(* Logix 5000 project; controller PLC_MCC1300_75F1 vendor 1 type 14 code 166 rev 32.11; software revision 32.04; part 6 of 83 *)
(* tags used below, declared in another part *)
   M352 : MAC_Conveyor;
   M353 : MAC_Conveyor;
   N14 : DINT[500];
   N30 : DINT[32];
   N31 : DINT[33];   // M2 to M4
   N32 : DINT[33];
   N40 : DINT[32];
   N7 : DINT[101];
   N802 : INT[420];
   N803 : INT[420];
   O : INT[128];
   T4 : TIMER[51];
   T47 : TIMER[32];

ADD_ON_INSTRUCTION GP_TrackingGetLength   (* revision 1.0 *)
VAR_IN_OUT
   INO_tLine : UDT_LINE_TRACKING; {required}
END_VAR
VAR_INPUT
   IN_StartConveyorIndex : DINT; {access None, required}
   IN_StopConveyorIndex : DINT; {access None, required}
END_VAR
VAR_OUTPUT
   OUT_dLength_cmm : DINT; {access None}
END_VAR
VAR
   TMP_dLineSize : DINT; {access None}
   TMP_dIndex : DINT; {access None}
END_VAR

ROUTINE Logic   (* structured text *)
   
   OUT_dLength_cmm := 0;
   size(INO_tLine.rgtTrkConv[0],0,TMP_dLineSize);
   IF IN_StartConveyorIndex >= 0 AND IN_StartConveyorIndex < TMP_dLineSize AND IN_StopConveyorIndex >= IN_StartConveyorIndex AND IN_StopConveyorIndex < TMP_dLineSize THEN
   	FOR TMP_dIndex := IN_StartConveyorIndex TO IN_StopConveyorIndex DO
   		OUT_dLength_cmm := OUT_dLength_cmm + INO_tLine.rgtTrkConv[TMP_dIndex].dLengthConveyor;
   	END_FOR;
   END_IF;
   
END_ROUTINE
END_ADD_ON_INSTRUCTION

ADD_ON_INSTRUCTION GP_TrackingPresencePlate   (* revision 1.0 *)
VAR_INPUT
   IN_dPositionStartSearch_cmm : DINT; {access None, required}   // Position of start searching plate
   IN_dPositionStopSearch_cmm : DINT; {access None, required}   // Position of stop searching plate
   IN_xConvoySearchSingle : BOOL; {access None, required}   // Search single cap in a convoy
END_VAR
VAR_IN_OUT
   INO_tLine : UDT_LINE_TRACKING; {required}   // Tracking area
END_VAR
VAR_OUTPUT
   OUT_xPlatePresence : BOOL; {access Read Only, required}
END_VAR
VAR
   TMP_dIndConv : DINT; {access None}
   TMP_dPositionMax_cmm : DINT; {access None}
   TMP_dPositionMin_cmm : DINT; {access None}
   TMP_dIndConvMax : DINT; {access None}
   TMP_dIndConvMin : DINT; {access None}
   TMP_dIndCap : DINT; {access None}
   TMP_dLineSize : DINT; {access None}
END_VAR

ROUTINE Logic   (* structured text *)
   
   OUT_xPlatePresence := 0;
   TMP_dPositionMax_cmm := IN_dPositionStopSearch_cmm;
   TMP_dPositionMin_cmm := IN_dPositionStartSearch_cmm;
   size(INO_tLine.rgtTrkConv[0],0,TMP_dLineSize);
   
   //Search The index of Conveyor
   FOR TMP_dIndConv := 0 TO TMP_dLineSize - 1 DO
       //Search Conveyor Index Min
       IF TMP_dPositionMin_cmm <= INO_tLine.rgtTrkConv[TMP_dIndConv].dEndPosition_cmm AND TMP_dPositionMin_cmm >= INO_tLine.rgtTrkConv[TMP_dIndConv].dStartPosition_cmm THEN
           TMP_dIndConvMin := TMP_dIndConv;
       END_IF;
       //Search Conveyor Index Max
       IF TMP_dPositionMax_cmm <= INO_tLine.rgtTrkConv[TMP_dIndConv].dEndPosition_cmm AND TMP_dPositionMax_cmm >= INO_tLine.rgtTrkConv[TMP_dIndConv].dStartPosition_cmm THEN
           TMP_dIndConvMax := TMP_dIndConv;
           EXIT;
       END_IF;
   END_FOR;
   
   FOR TMP_dIndConv := TMP_dIndConvMin TO TMP_dIndConvMax DO
       IF INO_tLine.rgtTrkConv[TMP_dIndConv].xGlassPresence THEN
           FOR TMP_dIndCap := 0 TO INO_tLine.rgtTrkConv[TMP_dIndConv].dIndexCaps DO
               OUT_xPlatePresence := (INO_tLine.rgtTrkConv[TMP_dIndConv].Cap[TMP_dIndCap].dPresenceHead_cmm >= TMP_dPositionMin_cmm
   			AND INO_tLine.rgtTrkConv[TMP_dIndConv].Cap[TMP_dIndCap].dPresenceHead_cmm <= TMP_dPositionMax_cmm)
               OR (INO_tLine.rgtTrkConv[TMP_dIndConv].Cap[TMP_dIndCap].dPresenceTail_cmm >= TMP_dPositionMin_cmm
   			AND INO_tLine.rgtTrkConv[TMP_dIndConv].Cap[TMP_dIndCap].dPresenceTail_cmm <= TMP_dPositionMax_cmm)
   			OR (INO_tLine.rgtTrkConv[TMP_dIndConv].Cap[TMP_dIndCap].dPresenceHead_cmm >= TMP_dPositionMax_cmm
   			AND INO_tLine.rgtTrkConv[TMP_dIndConv].Cap[TMP_dIndCap].dPresenceTail_cmm <= TMP_dPositionMin_cmm);
               IF OUT_xPlatePresence THEN
                   EXIT;
               END_IF;
           END_FOR;
       END_IF;
       IF OUT_xPlatePresence THEN
           EXIT;
       END_IF;
   END_FOR;
   
END_ROUTINE
END_ADD_ON_INSTRUCTION

ADD_ON_INSTRUCTION GP_TrackingSearchIDPlate   (* revision 1.0 *)
VAR_IN_OUT
   INO_tBufferPlate : UDT_LINE_BUFFER_PLATE; {required}
END_VAR
VAR_INPUT
   IN_dIDPlate : DINT; {access None, required}
END_VAR
VAR_OUTPUT
   OUT_dIndexPlate : DINT; {access None, required}
   OUT_xPlateIDFound : BOOL; {access Read Only, required}
END_VAR
VAR_IN_OUT
   INO_CONST_dMaxLites : DINT; {constant, required}
   INO_CONST_dMaxCaps : DINT; {constant, required}
END_VAR
VAR
   TMP_dInd : DINT; {access None}
   TMP_dLite : DINT; {access None}
   TMP_dCap : DINT; {access None}
   TMP_dBufferSize : DINT; {access None}
END_VAR

ROUTINE Logic   (* structured text *)
   
   size(INO_tBufferPlate.rgtPlate[0],0,TMP_dBufferSize);
   OUT_dIndexPlate := 0;//reset Output
   //Search Plate Index
   IF IN_dIDPlate <> 0 THEN
       FOR TMP_dInd := 0 TO TMP_dBufferSize - 1 DO
           FOR TMP_dCap := 0 TO INO_CONST_dMaxCaps - 1 DO
               FOR TMP_dLite := 0 TO INO_CONST_dMaxLites - 1 DO
   				IF INO_tBufferPlate.rgtPlate[TMP_dInd].tData.rgtCap[TMP_dCap].rgtLite[TMP_dLite].dID = IN_dIDPlate THEN
   					OUT_xPlateIDFound := 1;
   				END_IF;
                   IF OUT_xPlateIDFound THEN
                       OUT_dIndexPlate := TMP_dInd;//When found plate Exit from function
                       TND( );
                   END_IF;
               END_FOR;
           END_FOR;
       END_FOR;
   END_IF;
   
END_ROUTINE
END_ADD_ON_INSTRUCTION

ADD_ON_INSTRUCTION GP_TrackingSearchPlate   (* revision 1.0 *)
VAR_INPUT
   IN_dPositionStartSearch_cmm : DINT; {access None, required}   // Position of start searching plate
   IN_dPositionStopSearch_cmm : DINT; {access None, required}   // Position of stop searching plate
   IN_xConvoySearchSingle : BOOL; {access None, required}   // Search single cap in a convoy
END_VAR
VAR_IN_OUT
   INO_tLineTracking : UDT_LINE_TRACKING; {required}   // Tracking area
   INO_GP_SearchPlate : GP_TrackingSearchPlate_STC; {required}   // Search results
   INO_dNumOfConveyors : DINT; {constant, required}   // Number of conveyors in tracking area
   INO_dNumCapsConveyor : DINT; {constant, required}   // Max number of caps per conveyor
   INO_tLineBufferPlate : UDT_LINE_BUFFER_PLATE; {required}   // Buffer plate
END_VAR
VAR
   TMP_dIndConv : DINT; {access None}
   TMP_dPositionMax_cmm : DINT; {access None}
   TMP_dPositionMin_cmm : DINT; {access None}
   TMP_xStartGreater : BOOL; {access None}
   TMP_dIndConvMax : DINT; {access None}
   TMP_dIndConvMin : DINT; {access None}
   TMP_dIndCap : DINT; {access None}
   TMP_dHeadPos : DINT; {access None}
   TMP_DIndexOut : DINT; {access None}
   TMP_dLastPosHead_cmm : DINT; {access None}
   TMP_dLastPosTail_cmm : DINT; {access None}
   TMP_dTailPos : DINT; {access None}
   TMP_dPointerCap : DINT; {access None}
   TMP_dTailPointer : DINT; {access None}
   TMP_dHeadPointer : DINT; {access None}   // Head pointer
END_VAR

ROUTINE Logic   (* structured text *)
   
   //Start Greater of the END
   TMP_xStartGreater := IN_dPositionStartSearch_cmm >= IN_dPositionStopSearch_cmm;
   INO_GP_SearchPlate.xTailPresence := 0;
   INO_GP_SearchPlate.xHeadPresence := 0;
   
   FOR TMP_DIndexOut := 0 TO 4 DO
       INO_GP_SearchPlate.rgdHead_cmm[TMP_DIndexOut] := 0;
       INO_GP_SearchPlate.rgdTail_cmm[TMP_DIndexOut] := 0;
       INO_GP_SearchPlate.rgdHeadPointer[TMP_DIndexOut] := 0;
       INO_GP_SearchPlate.rgdTailPointer[TMP_DIndexOut] := 0;
       INO_GP_SearchPlate.rgxHead.[TMP_DIndexOut] := 0;
       INO_GP_SearchPlate.rgxTail.[TMP_DIndexOut] := 0;
   END_FOR;
   TMP_DIndexOut := 0;
   
   IF TMP_xStartGreater THEN
       TMP_dPositionMax_cmm := IN_dPositionStartSearch_cmm;
       TMP_dPositionMin_cmm := IN_dPositionStopSearch_cmm;
   ELSE
       TMP_dPositionMax_cmm := IN_dPositionStopSearch_cmm;
       TMP_dPositionMin_cmm := IN_dPositionStartSearch_cmm;
   END_IF;
   
   //Search The index of Conveyor
   FOR TMP_dIndConv := 0 TO INO_dNumOfConveyors - 1 DO
       //Search Conveyor Index Min
       IF  TMP_dPositionMin_cmm <= INO_tLineTracking.rgtTrkConv[TMP_dIndConv].dEndPosition_cmm
   		AND TMP_dPositionMin_cmm >= INO_tLineTracking.rgtTrkConv[TMP_dIndConv].dStartPosition_cmm THEN
           TMP_dIndConvMin := TMP_dIndConv;
       END_IF;
       //Search Conveyor Index Max
       IF TMP_dPositionMax_cmm <= INO_tLineTracking.rgtTrkConv[TMP_dIndConv].dEndPosition_cmm
   		AND TMP_dPositionMax_cmm >= INO_tLineTracking.rgtTrkConv[TMP_dIndConv].dStartPosition_cmm THEN
           TMP_dIndConvMax := TMP_dIndConv;
           EXIT;
       END_IF;
   END_FOR;
   
   IF TMP_xStartGreater THEN
       //Start To the Max
   
       TMP_dLastPosHead_cmm := TMP_dPositionMax_cmm+1;
       TMP_dLastPosTail_cmm := TMP_dPositionMax_cmm+1;
       FOR TMP_DIndexOut := 0 TO 4 DO
           TMP_dHeadPos := 0;
           TMP_dTailPos := 0;
           FOR TMP_dIndConv := TMP_dIndConvMax TO TMP_dIndConvMin BY -1 DO
               IF INO_tLineTracking.rgtTrkConv[TMP_dIndConv].xGlassPresence THEN
                   FOR TMP_dIndCap := 0 TO INO_tLineTracking.rgtTrkConv[TMP_dIndConv].dIndexCaps DO
   					IF TMP_dIndCap < INO_dNumCapsConveyor THEN //Check to avoid CPU fault in case of tracking errors
   	                    TMP_dPointerCap := INO_tLineTracking.rgtTrkConv[TMP_dIndConv].Cap[TMP_dIndCap].dPointer;
   	                    IF INO_tLineTracking.rgtTrkConv[TMP_dIndConv].Cap[TMP_dIndCap].dHeadPos_cmm >= TMP_dPositionMin_cmm
   	                        AND INO_tLineTracking.rgtTrkConv[TMP_dIndConv].Cap[TMP_dIndCap].dHeadPos_cmm <= TMP_dPositionMax_cmm
   							AND INO_tLineTracking.rgtTrkConv[TMP_dIndConv].Cap[TMP_dIndCap].dHeadPos_cmm >= TMP_dHeadPos
   	                        AND (INO_tLineBufferPlate.rgtPlate[TMP_dPointerCap].tTracking.dPreviousCapIndex <= 0 OR IN_xConvoySearchSingle)
   							AND INO_tLineTracking.rgtTrkConv[TMP_dIndConv].Cap[TMP_dIndCap].xHead
   	                        AND INO_tLineTracking.rgtTrkConv[TMP_dIndConv].Cap[TMP_dIndCap].dHeadPos_cmm < TMP_dLastPosHead_cmm
   	                        AND ((NOT INO_tLineBufferPlate.rgtPlate[TMP_dPointerCap].tTracking.xNotConsConvTrk)
   							OR TMP_dIndConv < INO_tLineBufferPlate.rgtPlate[TMP_dPointerCap].tTracking.dIndexConvNotCons) THEN
   	                        TMP_dHeadPos := INO_tLineTracking.rgtTrkConv[TMP_dIndConv].Cap[TMP_dIndCap].dHeadPos_cmm;
   	                        TMP_dHeadPointer := TMP_dPointerCap;
   	                    END_IF;
   
   	                    IF INO_tLineTracking.rgtTrkConv[TMP_dIndConv].Cap[TMP_dIndCap].dTailPos_cmm >= TMP_dPositionMin_cmm
   	                        AND INO_tLineTracking.rgtTrkConv[TMP_dIndConv].Cap[TMP_dIndCap].dTailPos_cmm <= TMP_dPositionMax_cmm
   							AND INO_tLineTracking.rgtTrkConv[TMP_dIndConv].Cap[TMP_dIndCap].dTailPos_cmm >= TMP_dTailPos
   	                        AND (INO_tLineBufferPlate.rgtPlate[TMP_dPointerCap].tTracking.dNextCapIndex <= 0
   							OR IN_xConvoySearchSingle) AND INO_tLineTracking.rgtTrkConv[TMP_dIndConv].Cap[TMP_dIndCap].xTail
   	                        AND INO_tLineTracking.rgtTrkConv[TMP_dIndConv].Cap[TMP_dIndCap].dTailPos_cmm < TMP_dLastPosTail_cmm
   	                        AND ((NOT INO_tLineBufferPlate.rgtPlate[TMP_dPointerCap].tTracking.xNotConsConvTrk)
   							OR TMP_dIndConv < INO_tLineBufferPlate.rgtPlate[TMP_dPointerCap].tTracking.dIndexConvNotCons) THEN
   	                        TMP_dTailPos := INO_tLineTracking.rgtTrkConv[TMP_dIndConv].Cap[TMP_dIndCap].dTailPos_cmm;
   	                        TMP_dTailPointer := TMP_dPointerCap;
   	                    END_IF;
   					END_IF;
                   END_FOR;
               END_IF;
           END_FOR;
           //Write Output
           IF TMP_dHeadPointer <> 0 THEN
               INO_GP_SearchPlate.rgdHead_cmm[TMP_DIndexOut] := TMP_dHeadPos;
               INO_GP_SearchPlate.rgdHeadPointer[TMP_DIndexOut] := TMP_dHeadPointer;
               INO_GP_SearchPlate.rgxHead.[TMP_DIndexOut] := 1;
               INO_GP_SearchPlate.xHeadPresence := 1;
               TMP_dLastPosHead_cmm := TMP_dHeadPos;
               TMP_dHeadPointer := 0;
           END_IF;
   
           IF TMP_dTailPointer <> 0 THEN
               INO_GP_SearchPlate.rgdTail_cmm[TMP_DIndexOut] := TMP_dTailPos;
               INO_GP_SearchPlate.rgdTailPointer[TMP_DIndexOut] := TMP_dTailPointer;
               INO_GP_SearchPlate.rgxTail.[TMP_DIndexOut] := 1;
               INO_GP_SearchPlate.xTailPresence := 1;
               TMP_dLastPosTail_cmm := TMP_dTailPos;
           END_IF;
   
           IF TMP_dTailPointer = 0 AND TMP_dHeadPointer = 0 THEN
               EXIT;
           END_IF;
           TMP_dTailPointer := 0;
           TMP_dHeadPointer := 0;
       END_FOR;
   
   ELSE
       TMP_dLastPosHead_cmm := TMP_dPositionMin_cmm - 1;
       TMP_dLastPosTail_cmm := TMP_dPositionMin_cmm - 1;
       //Start To the Min
       FOR TMP_DIndexOut := 0 TO 4 DO
           TMP_dHeadPos := TMP_dPositionMax_cmm;
           TMP_dTailPos := TMP_dPositionMax_cmm;
           FOR TMP_dIndConv := TMP_dIndConvMin TO TMP_dIndConvMax DO
   
               IF INO_tLineTracking.rgtTrkConv[TMP_dIndConv].xGlassPresence THEN
                   FOR TMP_dIndCap := 0 TO INO_tLineTracking.rgtTrkConv[TMP_dIndConv].dIndexCaps DO
   					IF TMP_dIndCap < INO_dNumCapsConveyor THEN // To avoid CPU fault in case of tracking error (too much caps in one conveyor)
   	                    TMP_dPointerCap := INO_tLineTracking.rgtTrkConv[TMP_dIndConv].Cap[TMP_dIndCap].dPointer;
   	                    IF INO_tLineTracking.rgtTrkConv[TMP_dIndConv].Cap[TMP_dIndCap].dHeadPos_cmm >= TMP_dPositionMin_cmm
   	                        AND INO_tLineTracking.rgtTrkConv[TMP_dIndConv].Cap[TMP_dIndCap].dHeadPos_cmm <= TMP_dPositionMax_cmm
   							AND INO_tLineTracking.rgtTrkConv[TMP_dIndConv].Cap[TMP_dIndCap].dHeadPos_cmm <= TMP_dHeadPos
   	                        AND (INO_tLineBufferPlate.rgtPlate[TMP_dPointerCap].tTracking.dPreviousCapIndex <= 0 OR IN_xConvoySearchSingle)
   							AND INO_tLineTracking.rgtTrkConv[TMP_dIndConv].Cap[TMP_dIndCap].xHead
   	                        AND INO_tLineTracking.rgtTrkConv[TMP_dIndConv].Cap[TMP_dIndCap].dHeadPos_cmm > TMP_dLastPosHead_cmm THEN
   	                        TMP_dHeadPos := INO_tLineTracking.rgtTrkConv[TMP_dIndConv].Cap[TMP_dIndCap].dHeadPos_cmm;
   	                        TMP_dHeadPointer := TMP_dPointerCap;
   	                    END_IF;
   
   	                    IF INO_tLineTracking.rgtTrkConv[TMP_dIndConv].Cap[TMP_dIndCap].dTailPos_cmm >= TMP_dPositionMin_cmm
   	                        AND INO_tLineTracking.rgtTrkConv[TMP_dIndConv].Cap[TMP_dIndCap].dTailPos_cmm <= TMP_dPositionMax_cmm
   							AND INO_tLineTracking.rgtTrkConv[TMP_dIndConv].Cap[TMP_dIndCap].dTailPos_cmm <= TMP_dTailPos
   	                        AND (INO_tLineBufferPlate.rgtPlate[TMP_dPointerCap].tTracking.dNextCapIndex <= 0 OR IN_xConvoySearchSingle)
   							AND INO_tLineTracking.rgtTrkConv[TMP_dIndConv].Cap[TMP_dIndCap].xTail
   	                        AND INO_tLineTracking.rgtTrkConv[TMP_dIndConv].Cap[TMP_dIndCap].dTailPos_cmm > TMP_dLastPosTail_cmm THEN
   	                        TMP_dTailPos := INO_tLineTracking.rgtTrkConv[TMP_dIndConv].Cap[TMP_dIndCap].dTailPos_cmm;
   	                        TMP_dTailPointer := TMP_dPointerCap;
   	                    END_IF;
   					END_IF;
   	            END_FOR;
               END_IF;
           END_FOR;
           //Write Output
           IF TMP_dHeadPointer <> 0 THEN
               INO_GP_SearchPlate.rgdHead_cmm[TMP_DIndexOut] := TMP_dHeadPos;
               INO_GP_SearchPlate.rgdHeadPointer[TMP_DIndexOut] := TMP_dHeadPointer;
               INO_GP_SearchPlate.rgxHead.[TMP_DIndexOut] := 1;
               INO_GP_SearchPlate.xHeadPresence := 1;
               TMP_dLastPosHead_cmm := TMP_dHeadPos;
               TMP_dHeadPointer := 0;
           END_IF;
   
           IF TMP_dTailPointer <> 0 THEN
               INO_GP_SearchPlate.rgdTail_cmm[TMP_DIndexOut] := TMP_dTailPos;
               INO_GP_SearchPlate.rgdTailPointer[TMP_DIndexOut] := TMP_dTailPointer;
               INO_GP_SearchPlate.rgxTail.[TMP_DIndexOut] := 1;
               INO_GP_SearchPlate.xTailPresence := 1;
               TMP_dLastPosTail_cmm := TMP_dTailPos;
           END_IF;
   
           IF TMP_dTailPointer = 0 AND TMP_dHeadPointer = 0 THEN
               EXIT;
           END_IF;
           TMP_dTailPointer := 0;
           TMP_dHeadPointer := 0;
       END_FOR;
   END_IF;
   
END_ROUTINE
END_ADD_ON_INSTRUCTION

ADD_ON_INSTRUCTION GP_TrackingValidateIndex   (* revision 1.0 *)
VAR_IN_OUT
   INO_tLineBufferPlate : UDT_LINE_BUFFER_PLATE; {required}   // Buffer Plate
   INO_dIDMemory : DINT; {required}   // Memory of ID
END_VAR
VAR_INPUT
   IN_dIndex : DINT; {access None, required}   // Index
END_VAR
VAR_OUTPUT
   OUT_xDataConsistance : BOOL; {access None, required}   // Data consistance
END_VAR

ROUTINE Logic   (* structured text *)
   
   IF IN_dIndex <> 0 THEN
   	IF INO_tLineBufferPlate.rgtPlate[IN_dIndex].tData.rgtCap[0].dID <> 0 AND (INO_tLineBufferPlate.rgtPlate[IN_dIndex].tData.rgtCap[0].dID = INO_dIDMemory OR INO_dIDMemory = 0) THEN
   		OUT_xDataConsistance := 1;
   	ELSE
   		OUT_xDataConsistance := 0;
   		INO_dIDMemory := 0;
   	END_IF;
   ELSE
   	INO_dIDMemory := 0;
   	OUT_xDataConsistance := 0;
   END_IF;
   
END_ROUTINE
END_ADD_ON_INSTRUCTION

VAR_GLOBAL   (* controller tags *)
   AUX_tBufferPlate_NULL : UDT_BufferPlate; {access Read Only}
   AUX_tCapsConveyor_NULL : UDT_CapsConveyor_ZC; {access Read Only}
   AUX_tConvoy_SL_NULL : UDT_Convoy_SL; {access Read Only}
   AUX_tConvoyCap_ZC_NULL : UDT_ConvoyCap_ZC; {access Read Only}
   AUX_tHMI_Lite_NULL : UDT_HMI_LITE; {access Read Only}
   AUX_xDebugNewPlate : BOOL; {access Read Only}
   AUX_xInitialize : BOOL; {access Read Only}
   Axies : MOTION_GROUP; {access Read Only}
   B102 : DINT[1];
   B107 : DINT[1];
   B112 : DINT[1];
   B117 : DINT[1];
   B122 : DINT[1];
   B127 : DINT[1];
   B132 : DINT[1];
   B151 : DINT[1];
   B152 : DINT[1];
   B153 : DINT[1];
   B154 : DINT[1];
   B155 : DINT[1];
   B156 : DINT[1];
   B157 : DINT[1];
   B158 : DINT[1];
   B159 : DINT[1];
   B160 : DINT[1];
   B161 : DINT[1];
   B162 : DINT[1];
   B163 : DINT[1];
   B164 : DINT[1];
   B165 : DINT[1];
   B166 : DINT[1];
   B167 : DINT[1];
   B168 : DINT[1];
   B169 : DINT[1];
   B170 : DINT[1];
   B171 : DINT[1];
   B172 : DINT[1];
   B175 : DINT[1];
   B176 : DINT[1] := ([0] := 2#0000_0000_0000_0000_0000_1100_0000_0000);
   B180 : DINT[10] := ([0] := 2#0000_0000_0000_0000_0001_1111_1001_0000, [1] := 2#0000_0000_0000_0000_0000_0000_0000_0001, [2] := 2#0000_0000_0000_0000_0001_0000_1011_0111, [4] := 2#0000_0000_0000_0000_0001_0000_0000_0000, [5] := 2#0000_0000_0000_0000_0000_0000_0011_0001, [6] := 2#0000_0000_0000_0000_1001_1110_0000_0000, [7] := 2#0000_0000_0000_0000_0001_0110_1101_1011, [9] := 2#0000_0000_0000_0000_0000_0000_1100_0000);
   B3 : DINT[51] := ([0] := 2#0000_0000_0000_0000_0010_0000_0000_0000, [1] := 2#0000_0000_0000_0000_0000_0000_1000_0000, [6] := 2#0000_0000_0000_0000_0000_0010_0000_0000, [7] := 2#0000_0000_0000_0000_1000_0000_0000_1000, [50] := 2#0000_0000_0000_0000_0000_0000_0001_0000);
        [0].0   // DUMMY for Red Stack lite
        [0].1   // VMCC M4 Mainline is Backed up Flush a CAP
        [10].14   // Always false Tony
        [10].15   // Tony test Bit
        [12].12   // M3CM04 Second. Trans. Conv 4 - Resync Photo-Eye North (Conveyor 4)
        [12].13   // M3CM05 Second. Trans. Conv 5 - Resync Photo-Eye North (Conveyor 5)
        [12].14   // M3CM06 Second. Trans. Conv 6 - Resync Photo-Eye North (Conveyor 6)
        [12].15   // M3CM07 Queue Conv 2 Resync Photo-Eye North (Conveyor 7)
        [13].0   // M3CM08 Queue Conv 3 Resync Photo-Eye North (Conveyor 8)
        [13].1   // M3CM08 Queue Conv 4 Resync Photo-Eye North (Conveyor 9)
        [13].2   // QUALITY SAMPLE XFER 201.010 Xfer Conv M3CM10 QC5 Resync PE North (Conveyor 10)
        [13].6   // TRANSFER 1A VHSC gating Photo-eye North
        [14].0   // Mainline is in Sleep Mode
        [14].1   // Mainline in Sleep Mode Stop Conveyors
        [14].2   // ink jet ons
        [14].3   // INK JET Cap needs Ink jet messg
        [14].4   // ink jet ons2
        [18].13   // TRANSFER 1 Oversize cap Photo-eye EAST
        [18].14   // TRANSFER 1 Oversize cap Photo-Eye WEST
        [18].15   // TRANSFER 1A Oversize cap Photo-eye EAST
        [19].0   // TRANSFER 1A Oversize cap Photo-Eye WEST
        [2].15   // M4 -->> M5 Cap information One shot
        [50].0   // Sample Shuttle Peg is Approaching
        [50].1   // Sample Shuttle Peg is Ready for Pick up
        [5].10   // VMCC 4 Drive Fault Has occurred
        [5].11   // VMCC 3 Drive fault Has occurred
        [6].10   // CONVEYOR 6 Resync Photo-Eye South M3CM06
        [6].11   // M3CM07 Queue Conv 2 Resync Photo-Eye South (Conveyor 7)
        [6].12   // M3CM08 Queue Conv 3 Resync Photo-Eye South (Conveyor 8)
        [6].13   // M3CM08 Queue Conv 4 Resync Photo-Eyes (Conveyor 9)
        [6].14   // QUALITY SAMPLE XFER 201.010 Xfer Conv M3CM10 QC 5 Resync PE South (Conveyor 10)
        [6].15   // M4CM04 Transfer 1 Resync Photo-Eye South (Conveyor 11)
        [6].8   // M3CM04 Second. Trans. Conv 4 - Resync Photo-Eye South (Conveyor 4)
        [6].9   // M3CM05 Second. Trans. Conv 5 - Resync Photo-Eye South (Conveyor 5)
        [7].0   // M4CM03 Transfer 1 Rolls B Resync Photo-Eye South (Conveyor 12)
        [7].1   // M4CM04 Transfer 1 Rolls C Resync Photo-Eye South (Conveyor 13)
        [7].2   // TRANSFER 1A VHSC gating Photo-eye South
        [7].3   // M4CM05 Transfer 1A Rolls A - Rsync Photo-Eye South (Conveyor 15)
        [7].4   // M4CM07 Transfer 1A Rolls B - Rsync Photo-Eye South (Conveyor 16)
        [7].5   // M4CM09 Transfer 1A Rolls C - Rsync Photo-Eye South (Conveyor 17)
   B41 : DINT[3] := ([2] := 2#0000_0000_0000_0000_1000_0000_0000_0000);
        [0].13   // Conveyor 13 Resync Window
        [0].14   // Conveyor 14 Resync Window
        [0].15   // Conveyor 15 Resync Window
        [0].2   // Conveyor 2 Resync Window
        [0].3   // Conveyor 3 Resync Window
        [0].4   // Conveyor 4 Resync Window
        [0].5   // Conveyor 5 Resync Window
        [0].6   // Conveyor 6 Resync Window
        [0].7   // Conveyor 7 Resync Window
        [0].8   // Conveyor 8 Resync Window
        [0].9   // Conveyor 9 Resync Window
        [1].0   // Conveyor 16 Resync Window
        [1].5   // Conveyor 21 Resync Window
        [1].6   // Conveyor 22 Resync Window
        [1].7   // Conveyor 23 Resync Window
        [1].8   // Conveyor 24 Resync Window
        [1].9   // Conveyor 25 Resync Window
        [2].0   // Conveyor 32 Resync Window
        [1].1   // Conveyor 17 Resync Window
        [1].10   // Conveyor 26 Resync Window
        [1].11   // Conveyor 27 Resync Window
        [1].12   // Conveyor 28 Resync Window
        [1].13   // Conveyor 29 Resync Window
        [1].14   // Conveyor 30 Resync Window
        [1].15   // Conveyor 31 Resync Window
        [1].2   // Conveyor 18 Resync Window
        [1].3   // Conveyor 19 Resync Window
        [1].4   // Conveyor 20 Resync Window
        [0].1   // Conveyor 1 Resync Window
        [0].10   // Conveyor 10 Resync Window
        [0].11   // Conveyor 11 Resync Window
        [0].12   // Conveyor 12 Resync Window
   B42 : DINT[3];
        [0].1   // Conveyor 1 Resync Input
        [0].10   // Conveyor 10 Resync Input
        [0].11   // Conveyor 11 Resync Input
        [0].12   // Conveyor 12 Resync Input
        [0].13   // Conveyor 13 Resync Input
        [0].14   // Conveyor 14 Resync Input
        [0].15   // Conveyor 15 Resync Input
        [0].2   // Conveyor 2 Resync Input
        [0].3   // Conveyor 3 Resync Input
        [0].4   // Conveyor 4 Resync Input
        [0].5   // Conveyor 5 Resync Input
        [0].6   // Conveyor 6 Resync Input
        [0].7   // Conveyor 7 Resync Input
        [0].8   // Conveyor 8 Resync Input
        [0].9   // Conveyor 9 Resync Input
        [1].0   // Conveyor 16 Resync Input
        [1].1   // Conveyor 17 Resync Input
        [1].10   // Conveyor 26 Resync Input
        [1].11   // Conveyor 27 Resync Input
        [1].12   // Conveyor 28 Resync Input
        [1].13   // Conveyor 29 Resync Input
        [1].14   // Conveyor 30 Resync Input
        [1].15   // Conveyor 31 Resync Input
        [1].2   // Conveyor 18 Resync Input
        [1].3   // Conveyor 19 Resync Input
        [1].4   // Conveyor 20 Resync Input
        [1].5   // Conveyor 21 Resync Input
        [1].6   // Conveyor 22 Resync Input
        [1].7   // Conveyor 23 Resync Input
        [1].8   // Conveyor 24 Resync Input
        [1].9   // Conveyor 25 Resync Input
        [2].0   // Conveyor 32 Resync Input
   B43 : DINT[3];
        [0].12   // Conveyor 12 Resync Output
        [0].13   // Conveyor 13 Resync Output
        [0].14   // Conveyor 14 Resync Output
        [0].15   // Conveyor 15 Resync Output
        [0].2   // Conveyor 2 Resync Output
        [0].3   // Conveyor 3 Resync Output
        [0].4   // Conveyor 4 Resync Output
        [0].5   // Conveyor 5 Resync Output
        [0].6   // Conveyor 6 Resync Output
        [0].7   // Conveyor 7 Resync Output
        [0].8   // Conveyor 8 Resync Output
        [0].9   // Conveyor 9 Resync Output
        [1].0   // Conveyor 16 Resync Output
        [1].1   // Conveyor 17 Resync Output
        [1].10   // Conveyor 26 Resync Output
        [1].11   // Conveyor 27 Resync Output
        [1].12   // Conveyor 28 Resync Output
        [1].13   // Conveyor 29 Resync Output
        [1].14   // Conveyor 30 Resync Output
        [1].15   // Conveyor 31 Resync Output
        [1].2   // Conveyor 18 Resync Output
        [1].3   // Conveyor 19 Resync Output
        [1].4   // Conveyor 20 Resync Output
        [1].5   // Conveyor 21 Resync Output
        [1].6   // Conveyor 22 Resync Output
        [1].7   // Conveyor 23 Resync Output
        [1].8   // Conveyor 24 Resync Output
        [1].9   // Conveyor 25 Resync Output
        [2].0   // Conveyor 32 Resync Output
        [0].1   // Conveyor 1 Resync Output
        [0].10   // Conveyor 10 Resync Output
        [0].11   // Conveyor 11 Resync Output
   B45 : DINT[3];
        [0].13   // Conveyor 13 Resync Input Leading Edge
        [0].14   // Conveyor 14 Resync Input Leading Edge
        [0].15   // Conveyor 15 Resync Input Leading Edge
        [0].2   // Conveyor 2 Resync Input Leading Edge
        [0].3   // Conveyor 3 Resync Input Leading Edge
        [0].4   // Conveyor 4 Resync Input Leading Edge
        [0].5   // Conveyor 5 Resync Input Leading Edge
        [0].6   // Conveyor 6 Resync Input Leading Edge
        [0].7   // Conveyor 7 Resync Input Leading Edge
        [0].8   // Conveyor 8 Resync Input Leading Edge
        [0].9   // Conveyor 9 Resync Input Leading Edge
        [1].0   // Conveyor 16 Resync Input Leading Edge
        [1].1   // Conveyor 17 Resync Input Leading Edge
        [1].10   // Conveyor 26 Resync Input Leading Edge
        [1].11   // Conveyor 27 Resync Input Leading Edge
        [1].12   // Conveyor 28 Resync Input Leading Edge
        [1].13   // Conveyor 29 Resync Input Leading Edge
        [1].14   // Conveyor 30 Resync Input Leading Edge
        [1].15   // Conveyor 31 Resync Input Leading Edge
        [1].2   // Conveyor 18 Resync Input Leading Edge
        [1].3   // Conveyor 19 Resync Input Leading Edge
        [1].4   // Conveyor 20 Resync Input Leading Edge
        [1].5   // Conveyor 21 Resync Input Leading Edge
        [1].6   // Conveyor 22 Resync Input Leading Edge
        [1].7   // Conveyor 23 Resync Input Leading Edge
        [1].8   // Conveyor 24 Resync Input Leading Edge
        [1].9   // Conveyor 25 Resync Input Leading Edge
        [2].0   // Conveyor 32 Resync Input Leading Edge
        [0].1   // Conveyor 1 Resync Input Leading Edge
        [0].10   // Conveyor 10 Resync Input Leading Edge
        [0].11   // Conveyor 11 Resync Input Leading Edge
        [0].12   // Conveyor 12 Resync Input Leading Edge
   B46 : DINT[3];
        [1].11   // Conveyor 27 Resync Input Trailing Edge
        [0].1   // Conveyor 1 Resync Input Trailing Edge
        [1].12   // Conveyor 28 Resync Input Trailing Edge
        [1].13   // Conveyor 29 Resync Input Trailing Edge
        [0].10   // Conveyor 10 Resync Input Trailing Edge
        [1].14   // Conveyor 30 Resync Input Trailing Edge
        [1].15   // Conveyor 31 Resync Input Trailing Edge
        [0].11   // Conveyor 11 Resync Input Trailing Edge
        [1].2   // Conveyor 18 Resync Input Trailing Edge
        [1].3   // Conveyor 19 Resync Input Trailing Edge
        [0].12   // Conveyor 12 Resync Input Trailing Edge
        [1].4   // Conveyor 20 Resync Input Trailing Edge
        [1].5   // Conveyor 21 Resync Input Trailing Edge
        [0].13   // Conveyor 13 Resync Input Trailing Edge
        [1].6   // Conveyor 22 Resync Input Trailing Edge
        [0].14   // Conveyor 14 Resync Input Trailing Edge
        [0].15   // Conveyor 15 Resync Input Trailing Edge
        [1].7   // Conveyor 23 Resync Input Trailing Edge
        [0].2   // Conveyor 2 Resync Input Trailing Edge
        [1].8   // Conveyor 24 Resync Input Trailing Edge
        [1].9   // Conveyor 25 Resync Input Trailing Edge
        [0].3   // Conveyor 3 Resync Input Trailing Edge
        [0].4   // Conveyor 4 Resync Input Trailing Edge
        [0].5   // Conveyor 5 Resync Input Trailing Edge
        [0].6   // Conveyor 6 Resync Input Trailing Edge
        [0].7   // Conveyor 7 Resync Input Trailing Edge
        [0].8   // Conveyor 8 Resync Input Trailing Edge
        [0].9   // Conveyor 9 Resync Input Trailing Edge
        [2].0   // Conveyor 32 Resync Input Trailing Edge
        [1].0   // Conveyor 16 Resync Input Trailing Edge
        [1].1   // Conveyor 17 Resync Input Trailing Edge
        [1].10   // Conveyor 26 Resync Input Trailing Edge
   B60 : DINT[4];
        [0].12   // Conveyor 12 Glass in Transit Bits
        [0].13   // Conveyor 13 Glass in Transit Bits
        [0].14   // Conveyor 14 Glass in Transit Bits
        [0].15   // Conveyor 15 Glass in Transit Bits
        [0].2   // Conveyor 2 Glass in Transit Bits
        [0].3   // Conveyor 3 Glass in Transit Bits
        [0].4   // Conveyor 4 Glass in Transit Bits
        [0].5   // Conveyor 5 Glass in Transit Bits
        [0].6   // Conveyor 6 Glass in Transit Bits
        [0].7   // Conveyor 7 Glass in Transit Bits
        [0].8   // Conveyor 8 Glass in Transit Bits
        [0].9   // Conveyor 9 Glass in Transit Bits
        [1].0   // Conveyor 16 Glass in Transit Bits
        [1].1   // Conveyor 17 Glass in Transit Bits
        [1].10   // Conveyor 26 Glass in Transit Bits
        [1].11   // Conveyor 27 Glass in Transit Bits
        [1].12   // Conveyor 28 Glass in Transit Bits
        [1].13   // Conveyor 29 Glass in Transit Bits
        [1].14   // Conveyor 30 Glass in Transit Bits
        [1].15   // Conveyor 31 Glass in Transit Bits
        [1].2   // Conveyor 18 Glass in Transit Bits
        [1].3   // Conveyor 19 Glass in Transit Bits
        [1].4   // Conveyor 20 Glass in Transit Bits
        [1].5   // Conveyor 21 Glass in Transit Bits
        [1].6   // Conveyor 22 Glass in Transit Bits
        [1].7   // Conveyor 23 Glass in Transit Bits
        [1].8   // Conveyor 24 Glass in Transit Bits
        [0].1   // Conveyor 1 Glass in Transit Bits
        [1].9   // Conveyor 25 Glass in Transit Bits
        [0].10   // Conveyor 10 Glass in Transit Bits
        [0].11   // Conveyor 11 Glass in Transit Bits
        [2].0   // Conveyor 32 Glass in Transit Bits
   B70 : DINT[13] := ([4] := 2#0000_0000_0000_0000_0000_0000_0000_0010, [6] := 2#0000_0000_0000_0000_0100_0000_0000_0000, [8] := 2#0000_0000_0000_0000_1101_0000_0000_1100);
        [0]   // TRANSFER 1 Status Bits
        [0].0   // TRANSFER 1 One conveyor transfer
        [0].1   // TRANSFER 1 Downstream half of transfer occuppied
        [0].2   // TRANSFER 1 Two conveyor Transfer
        [0].3   // TRANSFER 1 Downstream Total transfer Occupied
        [0].4   // TRANSFER 1 Three conveyor Transfer
        [0].5   // TRANSFER 1 Sample plate for Transfer 1
        [1].12   // TRANSFER 1 Upstream Cap is stopped at transfer
        [1].13   // TRANSFER 1 Downstream Cap is stopped at transfer
        [1].2   // TRANSFER 1 Lash Rolls A to Rolls B (i.e. force them to follow)
        [1].4   // TRANSFER 1 Upstream half of transfer Wait to see Gate input
        [1].5   // TRANSFER 1 Downstream half of transfer Wait to see Gate Input
        [1].8   // TRANSFER 1 Upstream half of Transfer VHSC Control Enabled
        [1].9   // TRANSFER 1 Downstream Half of Transfer VHSC Control Enabled
        [3].11   // TRANSFER 1 Leading cap Has exited xfer On upstream half only xfer
        [3].12   // TRANSFER 1 Trail edge Lock input
        [3].13   // TRANSFER 1 Conveyor is Seized for Transfer
        [4].0   // TRANSFER 1 Flush Signal
        [4].1   // TRANSFER 1 Setup Subroutine Glass Must Be Rotated before Packing
        [4].10   // TRANSFER 1 Rolls B Resync window Is a Two-Conv Transfer Cap
        [4].14   // TRANSFER 1 Glass was Aborted O/S
        [4].15   // TRANSFER 1 Occupied or Positioning a Cap
        [4].6   // TRANSFER 1 Transfer ABORTED!
        [4].7   // TRANSFER 1 Transfer is Complete
        [4].9   // TRANSFER 1 Stream 1 Size Matches the Jumbo Setup Size
        [5].1   // TRANSFER 1 Oversize cap Stopped at Transfer
        [5].15   // TRANSFER 1 Deck has been Raised manually
        [5].2   // TRANSFER 1 Glass is Ready for Transfer & No Vision Results Received when needed
        [5].3   // TRANSFER 1 Glass is Ready for Transfer & Vision Results were Received
        [6]   // TRANSFER 1 Transfer abort Reason History Bits
        [6].0   // Transfer abort Reason History Bit MANUAL ABORT
        [6].1   // REASON 1 Transfer Abort - Rack fault
        [6].10   // REASON 10 Transfer Abort - Deck raise Failure
        [6].11   // REASON 11 Transfer Abort - Duration Watchdog
        [6].12   // REASON 12 Transfer Abort - Size Mismatch
        [6].13   // REASON 13 Transfer Abort - Mainline Flush
        [6].14   // REASON 14 Transfer Abort - Transfer Disable Switch
        [6].15   // REASON 15 Transfer Abort - Mainline Vision Reject
        [6].2   // REASON 2 Transfer Abort - Leg equip. Failure
        [6].3   // REASON 3 Transfer Abort - Bad cap data To leg PLC
        [6].4   // REASON 4 Transfer Abort - Belt drive Fault
        [6].5   // REASON 5 Transfer Abort - LCR watchdog
        [6].6   // REASON 6 Transfer Abort - Rolls A Stop Watchdog
        [6].7   // REASON 7 Transfer Abort - Rolls B Stop Watchdog
        [6].8   // REASON 8 Transfer Abort - Rolls A Oversize cap
        [6].9   // REASON 9 Transfer Abort - Rolls B Oversize cap
        [7].0   // TRANSFER 1 One conveyor LCR
        [7].1   // TRANSFER 1 Downstream half Transfer LCR
        [7].2   // TRANSFER 1 Two conveyor LCR
        [7].3   // TRANSFER 1 Downstream Full Size Transfer LCR
        [7].4   // TRANSFER 1 Three conveyor LCR
        [8].0   // TRANSFER 1 Leading Cap Runout In Progress
        [8].1   // TRANSFER 1 Gap too small For one Conveyor Transfer
        [8].12   // TRANSFER 1 Conveyor 6 run permissives
        [8].13   // TRANSFER 1 Cap at Photo-Eye will Resync
        [8].15   // Valid data
        [8].2   // TRANSFER 1 Gap too small For two Conveyor Transfer
        [8].3   // TRANSFER 1 Gap too small For three Conveyor Transfer
        [8].4   // TRANSFER 1 Minimum gap For DECEL Is not Present!
        [9].0   // TRANSFER 1 Runout Sensors Checked OK Reset Warning Seal Circuit
        [9].1   // TRANSFER 1 Glass is Long enough to Reach the Center Runout Sensor
        [9].2   // TRANSFER 1 Glass is Long enough to Reach the West Runout Sensor
        [9].8   // TRANSFER 1 Cap is at Upstream QC PEs: Check for Take All
        [9].9   // TRANSFER 1 Cap at Upstream QC PEs Is a Known Vision System Reject
   BENCH_BUZZER : ALIAS FOR O[74].12;
   BENCH_MASTERUP : ALIAS FOR I[73].6;
   BT800_001 : MESSAGE;   // Block WRITE for M2CM1
        MessageParameters(ServiceCode := 16#004c, LocalElement := N802[0], ...)
   BT800_002 : MESSAGE;   // Block WRITE for M2CM2
        MessageParameters(ServiceCode := 16#004c, LocalElement := N802[20], ...)
   BT800_003 : MESSAGE;   // Block WRITE for M2CM3
        MessageParameters(ServiceCode := 16#004c, LocalElement := N802[40], ...)
   BT800_004 : MESSAGE;   // Block WRITE for M2CM4S
        MessageParameters(ServiceCode := 16#004c, LocalElement := N802[60], ...)
   BT800_005 : MESSAGE;   // Block WRITE for M2CM4N
        MessageParameters(ServiceCode := 16#004c, LocalElement := N802[80], ...)
   BT800_006 : MESSAGE;   // Block WRITE for M2CM5S
        MessageParameters(ServiceCode := 16#004c, LocalElement := N802[100], ...)
   BT800_007 : MESSAGE;   // Block WRITE for M2CM5N
        MessageParameters(ServiceCode := 16#004c, LocalElement := N802[120], ...)
   BT800_008 : MESSAGE;   // Block WRITE for M2CM6S
        MessageParameters(ServiceCode := 16#004c, LocalElement := N802[140], ...)
   BT800_009 : MESSAGE;   // Block WRITE for M2CM6N
        MessageParameters(ServiceCode := 16#004c, LocalElement := N802[160], ...)
   BT800_010 : MESSAGE;   // Block WRITE for M2CM7S
        MessageParameters(ServiceCode := 16#004c, LocalElement := N802[180], ...)
   BT800_011 : MESSAGE;   // Block WRITE for M2CM7N
        MessageParameters(ServiceCode := 16#004c, LocalElement := N802[200], ...)
   BT800_012 : MESSAGE;   // Block WRITE for M2CM8S
        MessageParameters(ServiceCode := 16#004c, LocalElement := N802[220], ...)
   BT800_013 : MESSAGE;   // Block WRITE for M2CM8N
        MessageParameters(ServiceCode := 16#004c, LocalElement := N802[240], ...)
   BT800_014 : MESSAGE;   // Block WRITE for M2CM9S
        MessageParameters(ServiceCode := 16#004c, LocalElement := N802[260], ...)
   BT800_015 : MESSAGE;   // Block WRITE for M2CM9N
        MessageParameters(ServiceCode := 16#004c, LocalElement := N802[280], ...)
   BT800_016 : MESSAGE;   // Block WRITE for M2CM10S
        MessageParameters(ServiceCode := 16#004c, LocalElement := N802[300], ...)
   BT800_017 : MESSAGE;   // Block WRITE for M2CM10N
        MessageParameters(ServiceCode := 16#004c, LocalElement := N802[320], ...)
   BT800_018 : MESSAGE;   // Block WRITE for M2CM11S
        MessageParameters(ServiceCode := 16#004c, LocalElement := N802[340], ...)
   BT800_019 : MESSAGE;   // Block WRITE for M2CM11N
        MessageParameters(ServiceCode := 16#004c, LocalElement := N802[360], ...)
   BT800_020 : MESSAGE;   // Block WRITE for M2CM12S
        MessageParameters(ServiceCode := 16#004c, LocalElement := N802[380], ...)
   BT800_021 : MESSAGE;   // Block Write for M2CM12N
        MessageParameters(ServiceCode := 16#004c, LocalElement := N802[400], ...)
   BT801_001 : MESSAGE;   // Block READ for M2CM01
        MessageParameters(ServiceCode := 16#004b, LocalElement := N803[0], ...)
   BT801_002 : MESSAGE;   // Block READ for M2CM2
        MessageParameters(ServiceCode := 16#004b, LocalElement := N803[20], ...)
   BT801_003 : MESSAGE;   // Block READ for M2CM3
        MessageParameters(ServiceCode := 16#004b, LocalElement := N803[40], ...)
   BT801_004 : MESSAGE;   // Block READ for M2CM4S
        MessageParameters(ServiceCode := 16#004b, LocalElement := N803[60], ...)
   BT801_005 : MESSAGE;   // Block READ for M2CM4N
        MessageParameters(ServiceCode := 16#004b, LocalElement := N803[80], ...)
   BT801_006 : MESSAGE;   // Block READ for M2CM5S
        MessageParameters(ServiceCode := 16#004b, LocalElement := N803[100], ...)
   BT801_007 : MESSAGE;   // Block READ for M2CM5N
        MessageParameters(ServiceCode := 16#004b, LocalElement := N803[120], ...)
   BT801_008 : MESSAGE;   // Block READ for M2CM6S
        MessageParameters(ServiceCode := 16#004b, LocalElement := N803[140], ...)
   BT801_009 : MESSAGE;   // Block READ for M2CM6N
        MessageParameters(ServiceCode := 16#004b, LocalElement := N803[160], ...)
   BT801_010 : MESSAGE;   // Block Read for M2CM7S
        MessageParameters(ServiceCode := 16#004b, LocalElement := N803[180], ...)
   BT801_011 : MESSAGE;   // Block Read for M2CM7N
        MessageParameters(ServiceCode := 16#004b, LocalElement := N803[200], ...)
   BT801_012 : MESSAGE;   // Block Read for M2CM8S
        MessageParameters(ServiceCode := 16#004b, LocalElement := N803[220], ...)
   BT801_013 : MESSAGE;   // Block Read for M2CM8N
        MessageParameters(ServiceCode := 16#004b, LocalElement := N803[240], ...)
   BT801_014 : MESSAGE;   // Block Read for M2CM9S
        MessageParameters(ServiceCode := 16#004b, LocalElement := N803[260], ...)
   BT801_015 : MESSAGE;   // Block Read for M2CM9N
        MessageParameters(ServiceCode := 16#004b, LocalElement := N803[280], ...)
   BT801_016 : MESSAGE;   // Block Read for M2CM10S
        MessageParameters(ServiceCode := 16#004b, LocalElement := N803[300], ...)
   BT801_017 : MESSAGE;   // Block Read for M2CM10N
        MessageParameters(ServiceCode := 16#004b, LocalElement := N803[320], ...)
   BT801_018 : MESSAGE;   // Block Read for M2CM11S
        MessageParameters(ServiceCode := 16#004b, LocalElement := N803[340], ...)
   BT801_019 : MESSAGE;   // Block Read for M2CM11N
        MessageParameters(ServiceCode := 16#004b, LocalElement := N803[360], ...)
   BT801_020 : MESSAGE;   // Block Read for M2CM12S
        MessageParameters(ServiceCode := 16#004b, LocalElement := N803[380], ...)
   BT801_021 : MESSAGE;   // Block Read for M2CM12N
        MessageParameters(ServiceCode := 16#004b, LocalElement := N803[400], ...)
   C104 : COUNTER[1];
   C109 : COUNTER[1];
   C114 : COUNTER[1];
   C119 : COUNTER[1];
   C124 : COUNTER[1];
   C129 : COUNTER[1] := ([0].PRE := 100);
   C134 : COUNTER[1];
   C183 : COUNTER[10] := ([0].PRE := 12, [0].CU := 1, [1].PRE := 3, [1].CU := 1, [2].PRE := 3, [2].CU := 1);
   C48 : COUNTER[101];
        [14]   // Conveyor 14 Lost Caps Counter
        [15]   // Conveyor 15 Lost Caps Counter
        [16]   // Conveyor 16 Lost Caps Counter
        [10]   // Conveyor 10 Lost Caps Counter
        [11]   // Conveyor 11 Lost Caps Counter
        [12]   // Conveyor 12 Lost Caps Counter
        [13]   // Conveyor 13 Lost Caps Counter
        [17]   // Conveyor 17 Lost Caps Counter
        [18]   // Conveyor 18 Lost Caps Counter
        [19]   // Conveyor 19 Lost Caps Counter
        [1]   // Conveyor 1 Lost Caps Counter
        [20]   // Conveyor 20 Lost Caps Counter
        [21]   // Conveyor 21 Lost Caps Counter
        [22]   // Conveyor 22 Lost Caps Counter
        [23]   // Conveyor 23 Lost Caps Counter
        [24]   // Conveyor 24 Lost Caps Counter
        [25]   // Conveyor 25 Lost Caps Counter
        [26]   // Conveyor 26 Lost Caps Counter
        [27]   // Conveyor 27 Lost Caps Counter
        [28]   // Conveyor 28 Lost Caps Counter
        [29]   // Conveyor 29 Lost Caps Counter
        [2]   // Conveyor 2 Lost Caps Counter
        [30]   // Conveyor 30 Lost Caps Counter
        [31]   // Conveyor 31 Lost Caps Counter
        [32]   // Conveyor 32 Lost Caps Counter
        [3]   // Conveyor 3 Lost Caps Counter
        [4]   // Conveyor 4 Lost Caps Counter
        [5]   // Conveyor 5 Lost Caps Counter
        [6]   // Conveyor 6 Lost Caps Counter
        [7]   // Conveyor 7 Lost Caps Counter
        [8]   // Conveyor 8 Lost Caps Counter
        [9]   // Conveyor 9 Lost Caps Counter
   C49 : COUNTER[33];
        [31]   // Conveyor 31 Resync window Tuning Counter
        [32]   // Conveyor 32 Resync window Tuning Counter
        [3]   // Conveyor 3 Resync window Tuning Counter
        [4]   // Conveyor 4 Resync window Tuning Counter
        [5]   // Conveyor 5 Resync window Tuning Counter
        [6]   // Conveyor 6 Resync window Tuning Counter
        [7]   // Conveyor 7 Resync window Tuning Counter
        [8]   // Conveyor 8 Resync window Tuning Counter
        [9]   // Conveyor 9 Resync window Tuning Counter
        [10]   // Conveyor 10 Resync window Tuning Counter
        [11]   // Conveyor 11 Resync window Tuning Counter
        [12]   // Conveyor 12 Resync window Tuning Counter
        [13]   // Conveyor 13 Resync window Tuning Counter
        [14]   // Conveyor 14 Resync window Tuning Counter
        [15]   // Conveyor 15 Resync window Tuning Counter
        [16]   // Conveyor 16 Resync window Tuning Counter
        [17]   // Conveyor 17 Resync window Tuning Counter
        [18]   // Conveyor 18 Resync window Tuning Counter
        [19]   // Conveyor 19 Resync window Tuning Counter
        [1]   // Conveyor 1 Resync window Tuning Counter
        [20]   // Conveyor 20 Resync window Tuning Counter
        [21]   // Conveyor 21 Resync window Tuning Counter
        [22]   // Conveyor 22 Resync window Tuning Counter
        [23]   // Conveyor 23 Resync window Tuning Counter
        [24]   // Conveyor 24 Resync window Tuning Counter
        [25]   // Conveyor 25 Resync window Tuning Counter
        [26]   // Conveyor 26 Resync window Tuning Counter
        [27]   // Conveyor 27 Resync window Tuning Counter
        [28]   // Conveyor 28 Resync window Tuning Counter
        [29]   // Conveyor 29 Resync window Tuning Counter
        [2]   // Conveyor 2 Resync window Tuning Counter
        [30]   // Conveyor 30 Resync window Tuning Counter
   C5 : COUNTER[51] := ([0].PRE := 10000, [0].ACC := 637, [1].PRE := 10000, [1].ACC := 573, [2].PRE := 10000, [2].ACC := 13, [3].PRE := 10000, [3].ACC := 546, [4].PRE := 1000, [4].ACC := 13, [5].PRE := 1000, [5].ACC := 541, [6].PRE := 1000, [6].ACC := 553, [7].PRE := 1000, [7].ACC := 563, [8].PRE := 1000, [8].ACC := 559, [9].PRE := 1000, [9].ACC := 551, [10].PRE := 1000, [10].ACC := 991, [11].PRE := 1000, [11].ACC := 545, [12].PRE := 10000, [12].ACC := 175, [13].PRE := 1000, [13].ACC := 549, [14].PRE := 1000, [14].ACC := 552, [15].PRE := 1000, [15].ACC := 547, [16].PRE := 10000, [16].ACC := 1164, [17].PRE := 1000, [17].ACC := 559, [18].PRE := 1000, [18].ACC := 550, [19].PRE := 1000, [19].ACC := 550, [20].PRE := 1000, [20].ACC := 545, [21].PRE := 1000, [21].ACC := 600, [22].PRE := 1000, [22].ACC := 601, [23].PRE := 1000, [23].ACC := 709, [25].PRE := 3, [25].ACC := 1, [30].PRE := 1000, [30].ACC := 60, [31].PRE := 1000, [31].ACC := 37, [32].PRE := 1000, [32].ACC := 52, [33].PRE := 1000, [33].ACC := 24, [34].PRE := 1000, [34].ACC := 166,
        [35].PRE := 1000, [35].ACC := 154, [36].PRE := 1000, [36].ACC := 121, [37].PRE := 1000, [37].ACC := 299, [38].PRE := 1000, [38].ACC := 8, [39].PRE := 1000, [39].ACC := 10, [40].PRE := 1000, [40].ACC := 418, [41].PRE := 1000, [41].ACC := 667, [42].PRE := 1000, [42].ACC := 251, [43].PRE := 10000, [43].ACC := 2936, [44].PRE := 10000, [44].ACC := 8, [45].PRE := 10000, [45].ACC := 1, [46].PRE := 10000, [46].ACC := 1, [50].PRE := 100, [50].ACC := 87);
        [20]   // TRIM DECK Fault Tracking: Number of Times M2CM12S Drive Faulted
        [2]   // TRIM DECK Fault Tracking: Number of Times M2CM03 Drive Faulted
        [3]   // TRIM DECK Fault Tracking: Number of Times M2CM04S Drive Faulted
        [4]   // TRIM DECK Fault Tracking: Number of Times M2CM05N Drive Faulted
        [17]   // TRIM DECK Fault Tracking: Number of Times M2CM09S Drive Faulted
        [13]   // TRIM DECK Fault Tracking: Number of Times M2CM05S Drive Faulted
        [21]   // Debug Counter Number of Times M2CM08 Drive Faulted
        [10]   // TRIM DECK Fault Tracking: Number of Times M2CM11N Drive Faulted
        [15]   // TRIM DECK Fault Tracking: Number of Times M2CM07N Drive Faulted
        [0]   // TRIM DECK Fault Tracking: Number of Times M2CM01 Drive Faulted
        [31]   // TRIM DECK Fault Tracking: Number of Times M2CM02 Drive is Stopped
        [32]   // TRIM DECK Fault Tracking: Number of Times M2CM03 Drive is Stopped
        [38]   // TRIM DECK Fault Tracking: Number of Times M2CM09 Drive is Stopped
        [6]   // TRIM DECK Fault Tracking: Number of Times M2CM07S Drive Faulted
        [7]   // TRIM DECK Fault Tracking: Number of Times M2CM08N Drive Faulted
        [33]   // TRIM DECK Fault Tracking: Number of Times M2CM04 Drive is Stopped
        [34]   // TRIM DECK Fault Tracking: Number of Times M2CM05 Drive is Stopped
        [35]   // TRIM DECK Fault Tracking: Number of Times M2CM06 Drive is Stopped
        [39]   // TRIM DECK Fault Tracking: Number of Times M2CM10 Drive is Stopped
        [8]   // TRIM DECK Fault Tracking: Number of Times M2CM09N Drive Faulted
        [40]   // TRIM DECK Fault Tracking: Number of Times M2CM11 Drive is Stopped
        [36]   // TRIM DECK Fault Tracking: Number of Times M2CM07 Drive is Stopped
        [41]   // TRIM DECK Fault Tracking: Number of Times M2CM12 Drive is Stopped
        [42]   // TRIM DECK Fault Tracking: Number of Times ANY Drive 1-6 is Stopped
        [9]   // TRIM DECK Fault Tracking: Number of Times M2CM10N Drive Faulted
        [37]   // TRIM DECK Fault Tracking: Number of Times M2CM08 Drive is Stopped
        [43]   // TRIM DECK Fault Tracking: Number of Times ANY Drive 7-12 is Stopped
        [5]   // TRIM DECK Fault Tracking: Number of Times M2CM06S Drive Faulted
        [16]   // TRIM DECK Fault Tracking: Number of Times M2CM08S Drive Faulted
        [50]   // M2 -->> MB Trim deck Drive system Critical Failure Count
        [14]   // TRIM DECK Fault Tracking: Number of Times M2CM06N Drive Faulted